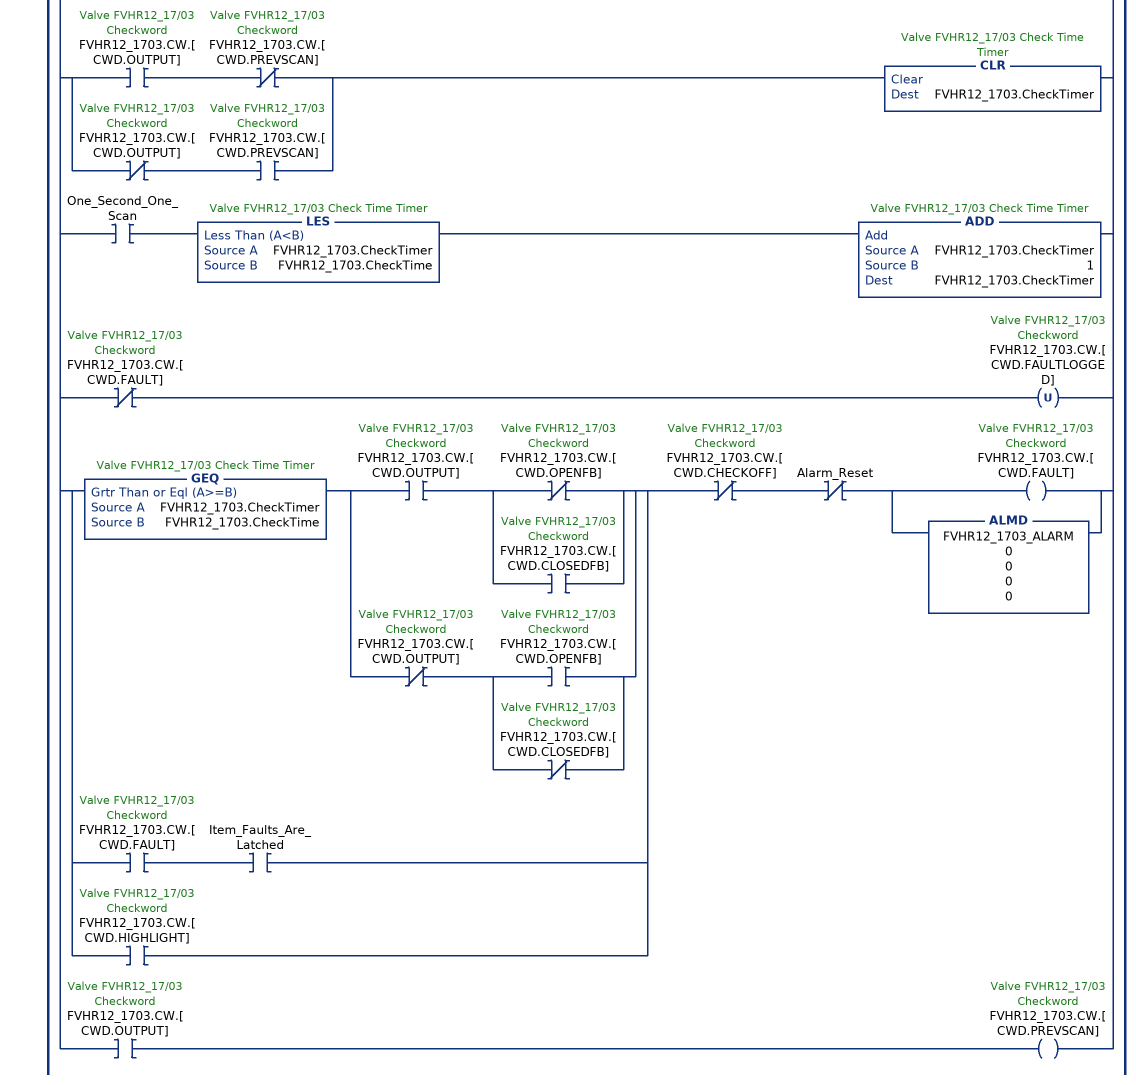
   71: [NEQ(FVHR12_1703.DriveBits,0) OTE(FVHR12_1703.CW.[CWD.AUTODRV]) ,[XIC(FVHR12_1703.CW.[CWD.AUTODRV]) XIO(FVHR12_1703.CW.[CWD.MANUAL]) ,XIC(FVHR12_1703.CW.[CWD.MANDRV]) XIC(FVHR12_1703.CW.[CWD.MANUAL]) ] OTE(FVHR12_1703.CW.[CWD.OUTPUT]) ,XIC(FVHR12_1703.CW.[CWD.OUTPUT]) OTE(FVHR12_1703_DR) ,XIC(S:FS) [OTU(FVHR12_1703.CW.[CWD.MANUAL]) ,LEQ(FVHR12_1703.CheckTime,0) MOV(Default_Check_Time,FVHR12_1703.CheckTime) ] ,[[XIC(FVHR12_1703_OP) XIO(Item_Simulation_Flag) ,XIC(Item_Simulation_Flag) XIC(FVHR12_1703.CW.[CWD.OUTPUT]) XIO(FVHR12_1703.CW.[CWD.SIMFAIL]) ] OTE(FVHR12_1703.CW.[CWD.OPENFB]) ,[XIC(FVHR12_1703_CL) XIO(Item_Simulation_Flag) ,XIC(Item_Simulation_Flag) XIO(FVHR12_1703.CW.[CWD.OUTPUT]) XIO(FVHR12_1703.CW.[CWD.SIMFAIL]) ] OTE(FVHR12_1703.CW.[CWD.CLOSEDFB]) ] ,[XIC(FVHR12_1703.CW.[CWD.OUTPUT]) XIO(FVHR12_1703.CW.[CWD.PREVSCAN]) ,XIO(FVHR12_1703.CW.[CWD.OUTPUT]) XIC(FVHR12_1703.CW.[CWD.PREVSCAN]) ] CLR(FVHR12_1703.CheckTimer) ,XIC(One_Second_One_Scan) LES(FVHR12_1703.CheckTimer,FVHR12_1703.CheckTime) ADD(FVHR12_1703.CheckTimer,1,FVHR12_1703.CheckTimer) ,XIO(FVHR12_1703.CW.[CWD.FAULT]) OTU(FVHR12_1703.CW.[CWD.FAULTLOGGED]) ,[GEQ(FVHR12_1703.CheckTimer,FVHR12_1703.CheckTime) [XIC(FVHR12_1703.CW.[CWD.OUTPUT]) [XIO(FVHR12_1703.CW.[CWD.OPENFB]) ,XIC(FVHR12_1703.CW.[CWD.CLOSEDFB]) ] ,XIO(FVHR12_1703.CW.[CWD.OUTPUT]) [XIC(FVHR12_1703.CW.[CWD.OPENFB]) ,XIO(FVHR12_1703.CW.[CWD.CLOSEDFB]) ] ] ,XIC(FVHR12_1703.CW.[CWD.FAULT]) XIC(Item_Faults_Are_Latched) ,XIC(FVHR12_1703.CW.[CWD.HIGHLIGHT]) ] XIO(FVHR12_1703.CW.[CWD.CHECKOFF]) XIO(Alarm_Reset) [OTE(FVHR12_1703.CW.[CWD.FAULT]) ,ALMD(FVHR12_1703_ALARM,0,0,0,0) ] ,XIC(FVHR12_1703.CW.[CWD.OUTPUT]) OTE(FVHR12_1703.CW.[CWD.PREVSCAN]) ];
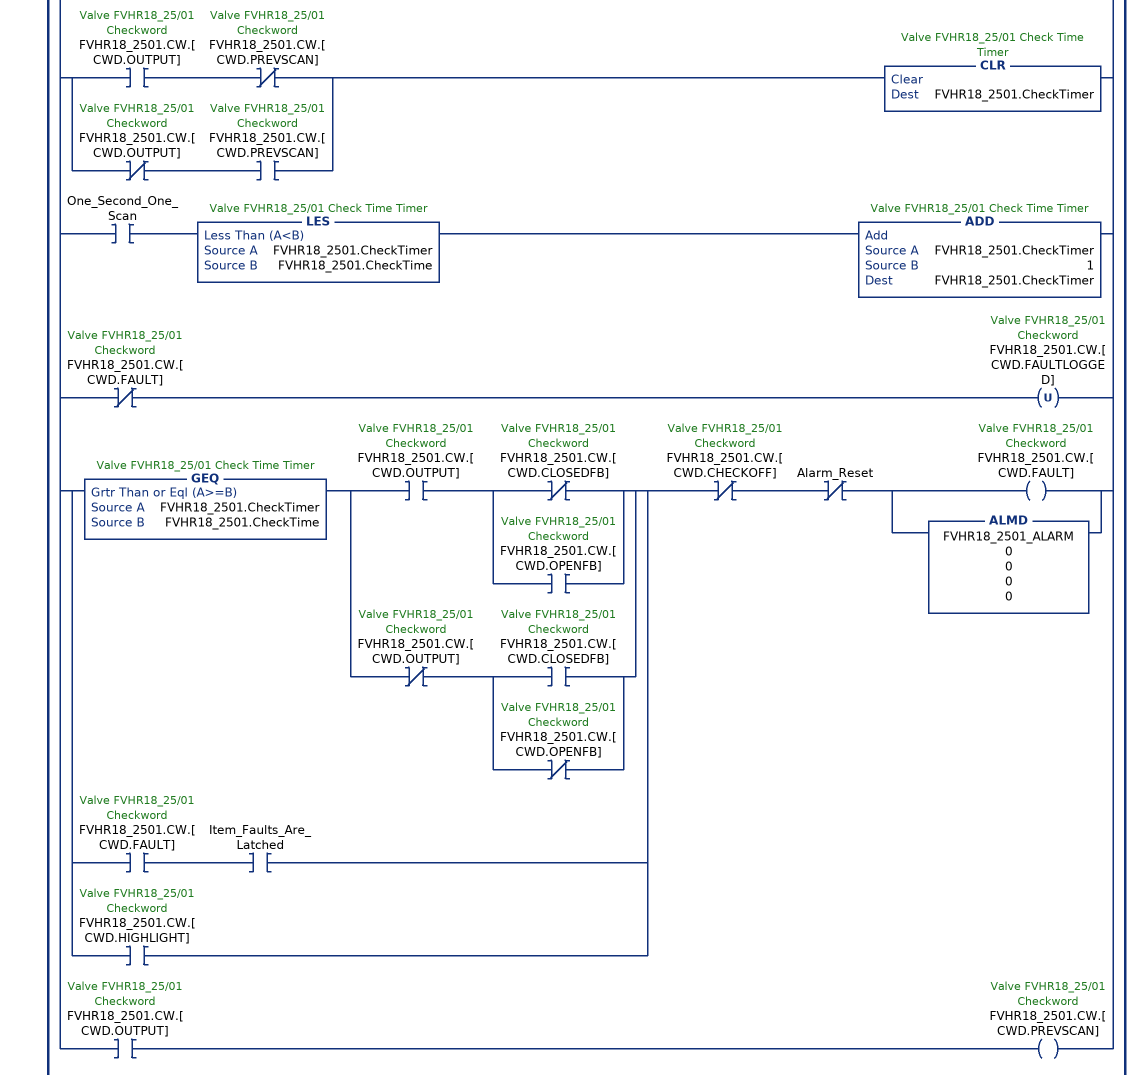
   72: [NEQ(FVHR18_2501.DriveBits,0) OTE(FVHR18_2501.CW.[CWD.AUTODRV]) ,[XIC(FVHR18_2501.CW.[CWD.AUTODRV]) XIO(FVHR18_2501.CW.[CWD.MANUAL]) ,XIC(FVHR18_2501.CW.[CWD.MANDRV]) XIC(FVHR18_2501.CW.[CWD.MANUAL]) ] OTE(FVHR18_2501.CW.[CWD.OUTPUT]) ,XIC(FVHR18_2501.CW.[CWD.OUTPUT]) OTE(FVHR18_2501_DR) ,XIC(S:FS) [OTU(FVHR18_2501.CW.[CWD.MANUAL]) ,LEQ(FVHR18_2501.CheckTime,0) MOV(Default_Check_Time,FVHR18_2501.CheckTime) ] ,[[XIC(FVHR18_2501_OP) XIO(Item_Simulation_Flag) ,XIC(Item_Simulation_Flag) XIC(FVHR18_2501.CW.[CWD.OUTPUT]) XIO(FVHR18_2501.CW.[CWD.SIMFAIL]) ] OTE(FVHR18_2501.CW.[CWD.OPENFB]) ,[XIC(FVHR18_2501_CL) XIO(Item_Simulation_Flag) ,XIC(Item_Simulation_Flag) XIO(FVHR18_2501.CW.[CWD.OUTPUT]) XIO(FVHR18_2501.CW.[CWD.SIMFAIL]) ] OTE(FVHR18_2501.CW.[CWD.CLOSEDFB]) ] ,[XIC(FVHR18_2501.CW.[CWD.OUTPUT]) XIO(FVHR18_2501.CW.[CWD.PREVSCAN]) ,XIO(FVHR18_2501.CW.[CWD.OUTPUT]) XIC(FVHR18_2501.CW.[CWD.PREVSCAN]) ] CLR(FVHR18_2501.CheckTimer) ,XIC(One_Second_One_Scan) LES(FVHR18_2501.CheckTimer,FVHR18_2501.CheckTime) ADD(FVHR18_2501.CheckTimer,1,FVHR18_2501.CheckTimer) ,XIO(FVHR18_2501.CW.[CWD.FAULT]) OTU(FVHR18_2501.CW.[CWD.FAULTLOGGED]) ,[GEQ(FVHR18_2501.CheckTimer,FVHR18_2501.CheckTime) [XIC(FVHR18_2501.CW.[CWD.OUTPUT]) [XIO(FVHR18_2501.CW.[CWD.CLOSEDFB]) ,XIC(FVHR18_2501.CW.[CWD.OPENFB]) ] ,XIO(FVHR18_2501.CW.[CWD.OUTPUT]) [XIC(FVHR18_2501.CW.[CWD.CLOSEDFB]) ,XIO(FVHR18_2501.CW.[CWD.OPENFB]) ] ] ,XIC(FVHR18_2501.CW.[CWD.FAULT]) XIC(Item_Faults_Are_Latched) ,XIC(FVHR18_2501.CW.[CWD.HIGHLIGHT]) ] XIO(FVHR18_2501.CW.[CWD.CHECKOFF]) XIO(Alarm_Reset) [OTE(FVHR18_2501.CW.[CWD.FAULT]) ,ALMD(FVHR18_2501_ALARM,0,0,0,0) ] ,XIC(FVHR18_2501.CW.[CWD.OUTPUT]) OTE(FVHR18_2501.CW.[CWD.PREVSCAN]) ];
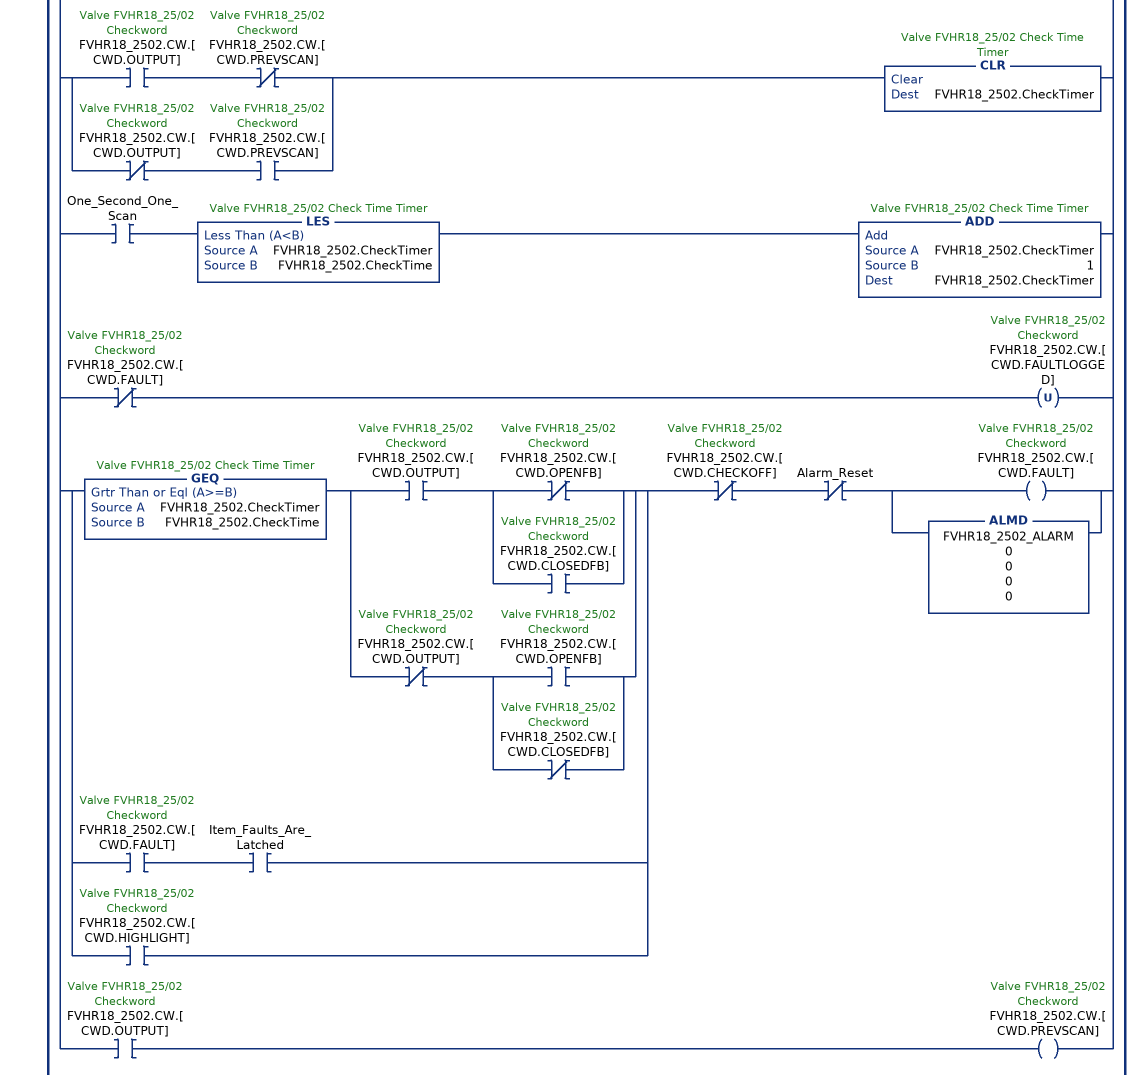
   73: [NEQ(FVHR18_2502.DriveBits,0) OTE(FVHR18_2502.CW.[CWD.AUTODRV]) ,[XIC(FVHR18_2502.CW.[CWD.AUTODRV]) XIO(FVHR18_2502.CW.[CWD.MANUAL]) ,XIC(FVHR18_2502.CW.[CWD.MANDRV]) XIC(FVHR18_2502.CW.[CWD.MANUAL]) ] OTE(FVHR18_2502.CW.[CWD.OUTPUT]) ,XIC(FVHR18_2502.CW.[CWD.OUTPUT]) OTE(FVHR18_2502_DR) ,XIC(S:FS) [OTU(FVHR18_2502.CW.[CWD.MANUAL]) ,LEQ(FVHR18_2502.CheckTime,0) MOV(Default_Check_Time,FVHR18_2502.CheckTime) ] ,[[XIC(FVHR18_2502_OP) XIO(Item_Simulation_Flag) ,XIC(Item_Simulation_Flag) XIC(FVHR18_2502.CW.[CWD.OUTPUT]) XIO(FVHR18_2502.CW.[CWD.SIMFAIL]) ] OTE(FVHR18_2502.CW.[CWD.OPENFB]) ,[XIC(FVHR18_2502_CL) XIO(Item_Simulation_Flag) ,XIC(Item_Simulation_Flag) XIO(FVHR18_2502.CW.[CWD.OUTPUT]) XIO(FVHR18_2502.CW.[CWD.SIMFAIL]) ] OTE(FVHR18_2502.CW.[CWD.CLOSEDFB]) ] ,[XIC(FVHR18_2502.CW.[CWD.OUTPUT]) XIO(FVHR18_2502.CW.[CWD.PREVSCAN]) ,XIO(FVHR18_2502.CW.[CWD.OUTPUT]) XIC(FVHR18_2502.CW.[CWD.PREVSCAN]) ] CLR(FVHR18_2502.CheckTimer) ,XIC(One_Second_One_Scan) LES(FVHR18_2502.CheckTimer,FVHR18_2502.CheckTime) ADD(FVHR18_2502.CheckTimer,1,FVHR18_2502.CheckTimer) ,XIO(FVHR18_2502.CW.[CWD.FAULT]) OTU(FVHR18_2502.CW.[CWD.FAULTLOGGED]) ,[GEQ(FVHR18_2502.CheckTimer,FVHR18_2502.CheckTime) [XIC(FVHR18_2502.CW.[CWD.OUTPUT]) [XIO(FVHR18_2502.CW.[CWD.OPENFB]) ,XIC(FVHR18_2502.CW.[CWD.CLOSEDFB]) ] ,XIO(FVHR18_2502.CW.[CWD.OUTPUT]) [XIC(FVHR18_2502.CW.[CWD.OPENFB]) ,XIO(FVHR18_2502.CW.[CWD.CLOSEDFB]) ] ] ,XIC(FVHR18_2502.CW.[CWD.FAULT]) XIC(Item_Faults_Are_Latched) ,XIC(FVHR18_2502.CW.[CWD.HIGHLIGHT]) ] XIO(FVHR18_2502.CW.[CWD.CHECKOFF]) XIO(Alarm_Reset) [OTE(FVHR18_2502.CW.[CWD.FAULT]) ,ALMD(FVHR18_2502_ALARM,0,0,0,0) ] ,XIC(FVHR18_2502.CW.[CWD.OUTPUT]) OTE(FVHR18_2502.CW.[CWD.PREVSCAN]) ];
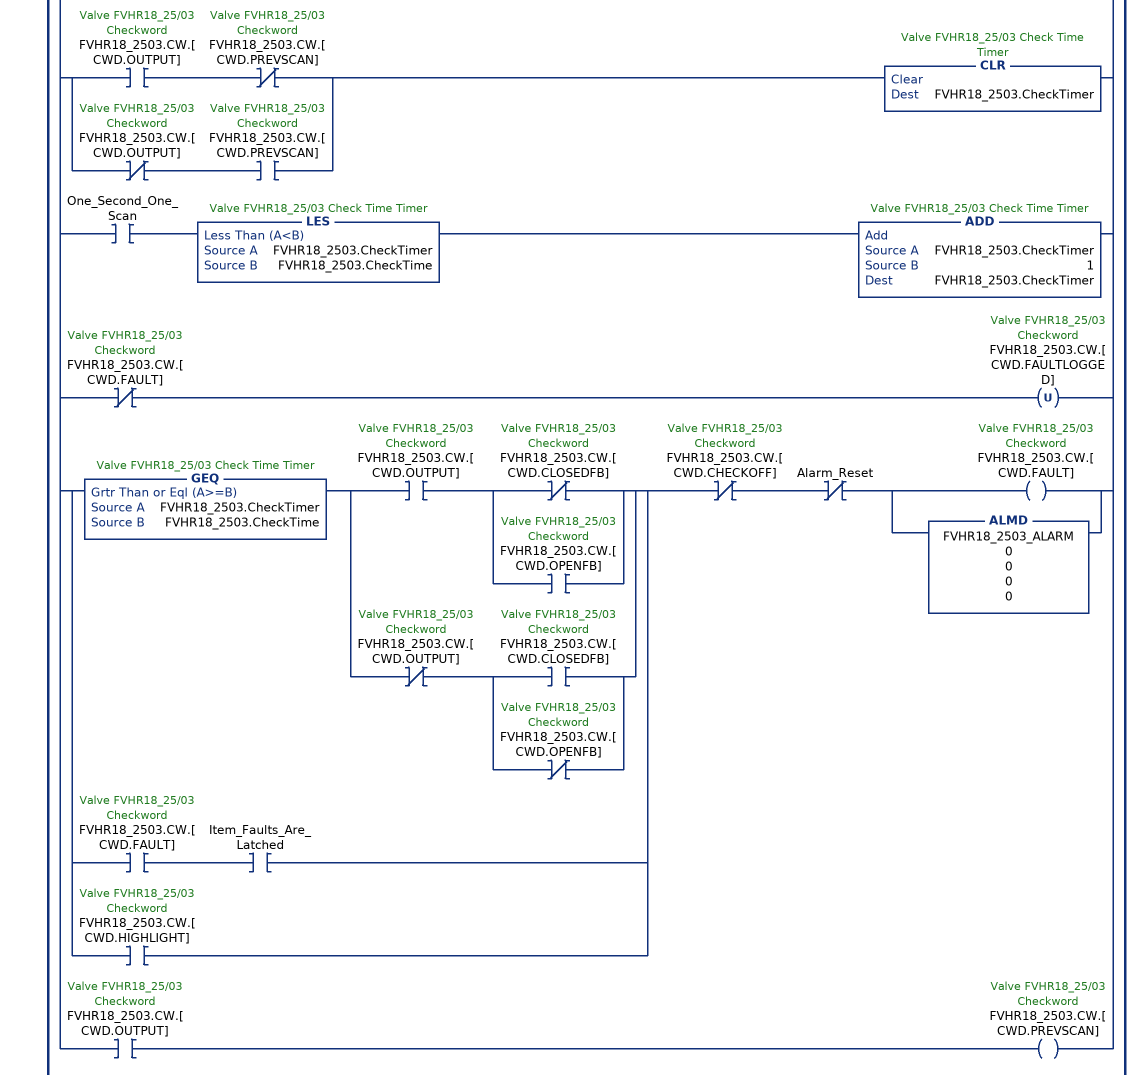
   74: [NEQ(FVHR18_2503.DriveBits,0) OTE(FVHR18_2503.CW.[CWD.AUTODRV]) ,[XIC(FVHR18_2503.CW.[CWD.AUTODRV]) XIO(FVHR18_2503.CW.[CWD.MANUAL]) ,XIC(FVHR18_2503.CW.[CWD.MANDRV]) XIC(FVHR18_2503.CW.[CWD.MANUAL]) ] OTE(FVHR18_2503.CW.[CWD.OUTPUT]) ,XIC(FVHR18_2503.CW.[CWD.OUTPUT]) OTE(FVHR18_2503_DR) ,XIC(S:FS) [OTU(FVHR18_2503.CW.[CWD.MANUAL]) ,LEQ(FVHR18_2503.CheckTime,0) MOV(Default_Check_Time,FVHR18_2503.CheckTime) ] ,[[XIC(FVHR18_2503_OP) XIO(Item_Simulation_Flag) ,XIC(Item_Simulation_Flag) XIC(FVHR18_2503.CW.[CWD.OUTPUT]) XIO(FVHR18_2503.CW.[CWD.SIMFAIL]) ] OTE(FVHR18_2503.CW.[CWD.OPENFB]) ,[XIC(FVHR18_2503_CL) XIO(Item_Simulation_Flag) ,XIC(Item_Simulation_Flag) XIO(FVHR18_2503.CW.[CWD.OUTPUT]) XIO(FVHR18_2503.CW.[CWD.SIMFAIL]) ] OTE(FVHR18_2503.CW.[CWD.CLOSEDFB]) ] ,[XIC(FVHR18_2503.CW.[CWD.OUTPUT]) XIO(FVHR18_2503.CW.[CWD.PREVSCAN]) ,XIO(FVHR18_2503.CW.[CWD.OUTPUT]) XIC(FVHR18_2503.CW.[CWD.PREVSCAN]) ] CLR(FVHR18_2503.CheckTimer) ,XIC(One_Second_One_Scan) LES(FVHR18_2503.CheckTimer,FVHR18_2503.CheckTime) ADD(FVHR18_2503.CheckTimer,1,FVHR18_2503.CheckTimer) ,XIO(FVHR18_2503.CW.[CWD.FAULT]) OTU(FVHR18_2503.CW.[CWD.FAULTLOGGED]) ,[GEQ(FVHR18_2503.CheckTimer,FVHR18_2503.CheckTime) [XIC(FVHR18_2503.CW.[CWD.OUTPUT]) [XIO(FVHR18_2503.CW.[CWD.CLOSEDFB]) ,XIC(FVHR18_2503.CW.[CWD.OPENFB]) ] ,XIO(FVHR18_2503.CW.[CWD.OUTPUT]) [XIC(FVHR18_2503.CW.[CWD.CLOSEDFB]) ,XIO(FVHR18_2503.CW.[CWD.OPENFB]) ] ] ,XIC(FVHR18_2503.CW.[CWD.FAULT]) XIC(Item_Faults_Are_Latched) ,XIC(FVHR18_2503.CW.[CWD.HIGHLIGHT]) ] XIO(FVHR18_2503.CW.[CWD.CHECKOFF]) XIO(Alarm_Reset) [OTE(FVHR18_2503.CW.[CWD.FAULT]) ,ALMD(FVHR18_2503_ALARM,0,0,0,0) ] ,XIC(FVHR18_2503.CW.[CWD.OUTPUT]) OTE(FVHR18_2503.CW.[CWD.PREVSCAN]) ];
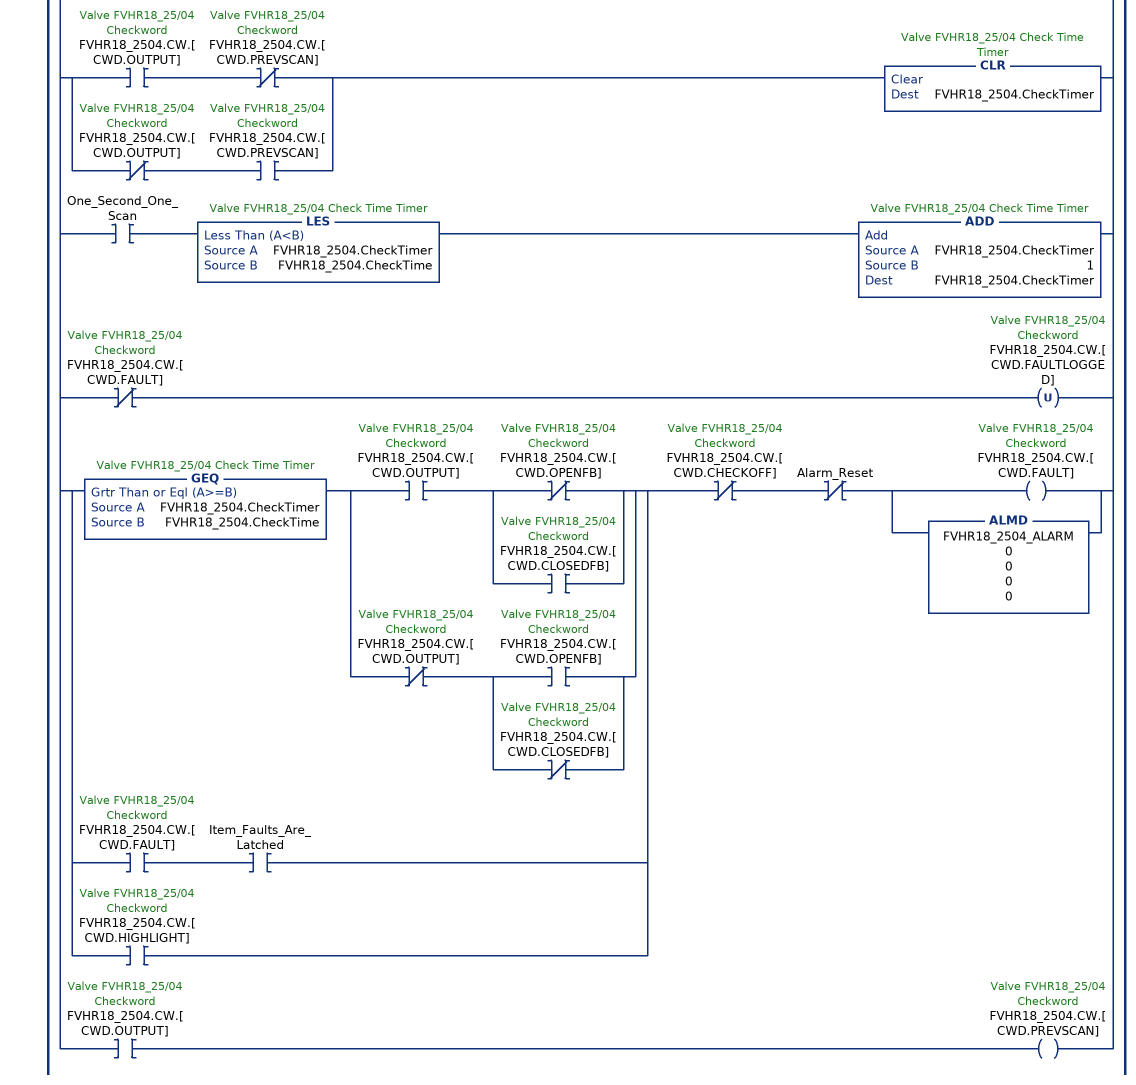
   75: [NEQ(FVHR18_2504.DriveBits,0) OTE(FVHR18_2504.CW.[CWD.AUTODRV]) ,[XIC(FVHR18_2504.CW.[CWD.AUTODRV]) XIO(FVHR18_2504.CW.[CWD.MANUAL]) ,XIC(FVHR18_2504.CW.[CWD.MANDRV]) XIC(FVHR18_2504.CW.[CWD.MANUAL]) ] OTE(FVHR18_2504.CW.[CWD.OUTPUT]) ,XIC(FVHR18_2504.CW.[CWD.OUTPUT]) OTE(FVHR18_2504_DR) ,XIC(S:FS) [OTU(FVHR18_2504.CW.[CWD.MANUAL]) ,LEQ(FVHR18_2504.CheckTime,0) MOV(Default_Check_Time,FVHR18_2504.CheckTime) ] ,[[XIC(FVHR18_2504_OP) XIO(Item_Simulation_Flag) ,XIC(Item_Simulation_Flag) XIC(FVHR18_2504.CW.[CWD.OUTPUT]) XIO(FVHR18_2504.CW.[CWD.SIMFAIL]) ] OTE(FVHR18_2504.CW.[CWD.OPENFB]) ,[XIC(FVHR18_2504_CL) XIO(Item_Simulation_Flag) ,XIC(Item_Simulation_Flag) XIO(FVHR18_2504.CW.[CWD.OUTPUT]) XIO(FVHR18_2504.CW.[CWD.SIMFAIL]) ] OTE(FVHR18_2504.CW.[CWD.CLOSEDFB]) ] ,[XIC(FVHR18_2504.CW.[CWD.OUTPUT]) XIO(FVHR18_2504.CW.[CWD.PREVSCAN]) ,XIO(FVHR18_2504.CW.[CWD.OUTPUT]) XIC(FVHR18_2504.CW.[CWD.PREVSCAN]) ] CLR(FVHR18_2504.CheckTimer) ,XIC(One_Second_One_Scan) LES(FVHR18_2504.CheckTimer,FVHR18_2504.CheckTime) ADD(FVHR18_2504.CheckTimer,1,FVHR18_2504.CheckTimer) ,XIO(FVHR18_2504.CW.[CWD.FAULT]) OTU(FVHR18_2504.CW.[CWD.FAULTLOGGED]) ,[GEQ(FVHR18_2504.CheckTimer,FVHR18_2504.CheckTime) [XIC(FVHR18_2504.CW.[CWD.OUTPUT]) [XIO(FVHR18_2504.CW.[CWD.OPENFB]) ,XIC(FVHR18_2504.CW.[CWD.CLOSEDFB]) ] ,XIO(FVHR18_2504.CW.[CWD.OUTPUT]) [XIC(FVHR18_2504.CW.[CWD.OPENFB]) ,XIO(FVHR18_2504.CW.[CWD.CLOSEDFB]) ] ] ,XIC(FVHR18_2504.CW.[CWD.FAULT]) XIC(Item_Faults_Are_Latched) ,XIC(FVHR18_2504.CW.[CWD.HIGHLIGHT]) ] XIO(FVHR18_2504.CW.[CWD.CHECKOFF]) XIO(Alarm_Reset) [OTE(FVHR18_2504.CW.[CWD.FAULT]) ,ALMD(FVHR18_2504_ALARM,0,0,0,0) ] ,XIC(FVHR18_2504.CW.[CWD.OUTPUT]) OTE(FVHR18_2504.CW.[CWD.PREVSCAN]) ];
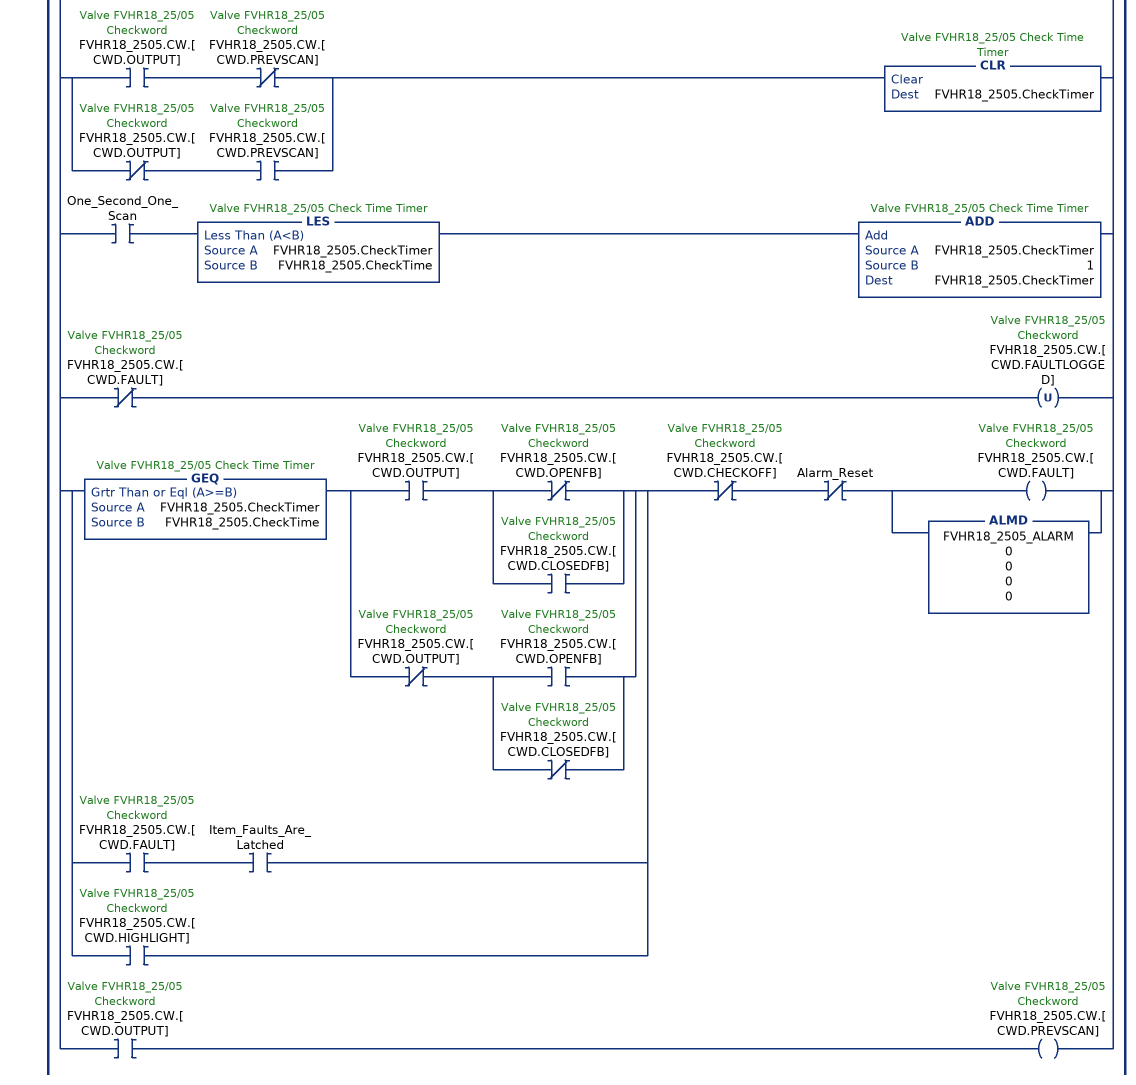
   76: [NEQ(FVHR18_2505.DriveBits,0) OTE(FVHR18_2505.CW.[CWD.AUTODRV]) ,[XIC(FVHR18_2505.CW.[CWD.AUTODRV]) XIO(FVHR18_2505.CW.[CWD.MANUAL]) ,XIC(FVHR18_2505.CW.[CWD.MANDRV]) XIC(FVHR18_2505.CW.[CWD.MANUAL]) ] OTE(FVHR18_2505.CW.[CWD.OUTPUT]) ,XIC(FVHR18_2505.CW.[CWD.OUTPUT]) OTE(FVHR18_2505_DR) ,XIC(S:FS) [OTU(FVHR18_2505.CW.[CWD.MANUAL]) ,LEQ(FVHR18_2505.CheckTime,0) MOV(Default_Check_Time,FVHR18_2505.CheckTime) ] ,[[XIC(FVHR18_2505_OP) XIO(Item_Simulation_Flag) ,XIC(Item_Simulation_Flag) XIC(FVHR18_2505.CW.[CWD.OUTPUT]) XIO(FVHR18_2505.CW.[CWD.SIMFAIL]) ] OTE(FVHR18_2505.CW.[CWD.OPENFB]) ,[XIC(FVHR18_2505_CL) XIO(Item_Simulation_Flag) ,XIC(Item_Simulation_Flag) XIO(FVHR18_2505.CW.[CWD.OUTPUT]) XIO(FVHR18_2505.CW.[CWD.SIMFAIL]) ] OTE(FVHR18_2505.CW.[CWD.CLOSEDFB]) ] ,[XIC(FVHR18_2505.CW.[CWD.OUTPUT]) XIO(FVHR18_2505.CW.[CWD.PREVSCAN]) ,XIO(FVHR18_2505.CW.[CWD.OUTPUT]) XIC(FVHR18_2505.CW.[CWD.PREVSCAN]) ] CLR(FVHR18_2505.CheckTimer) ,XIC(One_Second_One_Scan) LES(FVHR18_2505.CheckTimer,FVHR18_2505.CheckTime) ADD(FVHR18_2505.CheckTimer,1,FVHR18_2505.CheckTimer) ,XIO(FVHR18_2505.CW.[CWD.FAULT]) OTU(FVHR18_2505.CW.[CWD.FAULTLOGGED]) ,[GEQ(FVHR18_2505.CheckTimer,FVHR18_2505.CheckTime) [XIC(FVHR18_2505.CW.[CWD.OUTPUT]) [XIO(FVHR18_2505.CW.[CWD.OPENFB]) ,XIC(FVHR18_2505.CW.[CWD.CLOSEDFB]) ] ,XIO(FVHR18_2505.CW.[CWD.OUTPUT]) [XIC(FVHR18_2505.CW.[CWD.OPENFB]) ,XIO(FVHR18_2505.CW.[CWD.CLOSEDFB]) ] ] ,XIC(FVHR18_2505.CW.[CWD.FAULT]) XIC(Item_Faults_Are_Latched) ,XIC(FVHR18_2505.CW.[CWD.HIGHLIGHT]) ] XIO(FVHR18_2505.CW.[CWD.CHECKOFF]) XIO(Alarm_Reset) [OTE(FVHR18_2505.CW.[CWD.FAULT]) ,ALMD(FVHR18_2505_ALARM,0,0,0,0) ] ,XIC(FVHR18_2505.CW.[CWD.OUTPUT]) OTE(FVHR18_2505.CW.[CWD.PREVSCAN]) ];
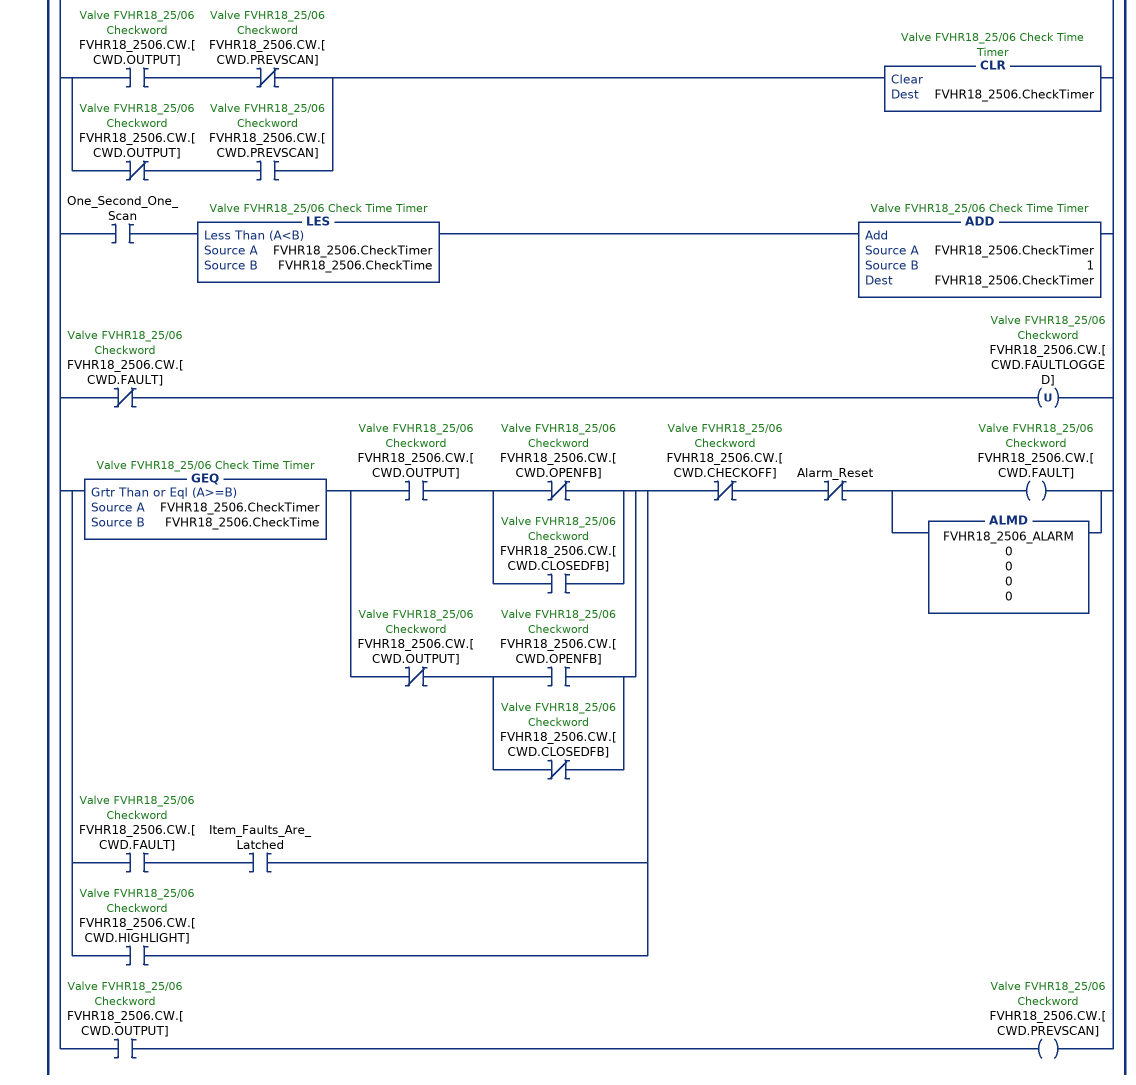
   77: [NEQ(FVHR18_2506.DriveBits,0) OTE(FVHR18_2506.CW.[CWD.AUTODRV]) ,[XIC(FVHR18_2506.CW.[CWD.AUTODRV]) XIO(FVHR18_2506.CW.[CWD.MANUAL]) ,XIC(FVHR18_2506.CW.[CWD.MANDRV]) XIC(FVHR18_2506.CW.[CWD.MANUAL]) ] OTE(FVHR18_2506.CW.[CWD.OUTPUT]) ,XIC(FVHR18_2506.CW.[CWD.OUTPUT]) OTE(FVHR18_2506_DR) ,XIC(S:FS) [OTU(FVHR18_2506.CW.[CWD.MANUAL]) ,LEQ(FVHR18_2506.CheckTime,0) MOV(Default_Check_Time,FVHR18_2506.CheckTime) ] ,[[XIC(FVHR18_2506_OP) XIO(Item_Simulation_Flag) ,XIC(Item_Simulation_Flag) XIC(FVHR18_2506.CW.[CWD.OUTPUT]) XIO(FVHR18_2506.CW.[CWD.SIMFAIL]) ] OTE(FVHR18_2506.CW.[CWD.OPENFB]) ,[XIC(FVHR18_2506_CL) XIO(Item_Simulation_Flag) ,XIC(Item_Simulation_Flag) XIO(FVHR18_2506.CW.[CWD.OUTPUT]) XIO(FVHR18_2506.CW.[CWD.SIMFAIL]) ] OTE(FVHR18_2506.CW.[CWD.CLOSEDFB]) ] ,[XIC(FVHR18_2506.CW.[CWD.OUTPUT]) XIO(FVHR18_2506.CW.[CWD.PREVSCAN]) ,XIO(FVHR18_2506.CW.[CWD.OUTPUT]) XIC(FVHR18_2506.CW.[CWD.PREVSCAN]) ] CLR(FVHR18_2506.CheckTimer) ,XIC(One_Second_One_Scan) LES(FVHR18_2506.CheckTimer,FVHR18_2506.CheckTime) ADD(FVHR18_2506.CheckTimer,1,FVHR18_2506.CheckTimer) ,XIO(FVHR18_2506.CW.[CWD.FAULT]) OTU(FVHR18_2506.CW.[CWD.FAULTLOGGED]) ,[GEQ(FVHR18_2506.CheckTimer,FVHR18_2506.CheckTime) [XIC(FVHR18_2506.CW.[CWD.OUTPUT]) [XIO(FVHR18_2506.CW.[CWD.OPENFB]) ,XIC(FVHR18_2506.CW.[CWD.CLOSEDFB]) ] ,XIO(FVHR18_2506.CW.[CWD.OUTPUT]) [XIC(FVHR18_2506.CW.[CWD.OPENFB]) ,XIO(FVHR18_2506.CW.[CWD.CLOSEDFB]) ] ] ,XIC(FVHR18_2506.CW.[CWD.FAULT]) XIC(Item_Faults_Are_Latched) ,XIC(FVHR18_2506.CW.[CWD.HIGHLIGHT]) ] XIO(FVHR18_2506.CW.[CWD.CHECKOFF]) XIO(Alarm_Reset) [OTE(FVHR18_2506.CW.[CWD.FAULT]) ,ALMD(FVHR18_2506_ALARM,0,0,0,0) ] ,XIC(FVHR18_2506.CW.[CWD.OUTPUT]) OTE(FVHR18_2506.CW.[CWD.PREVSCAN]) ];
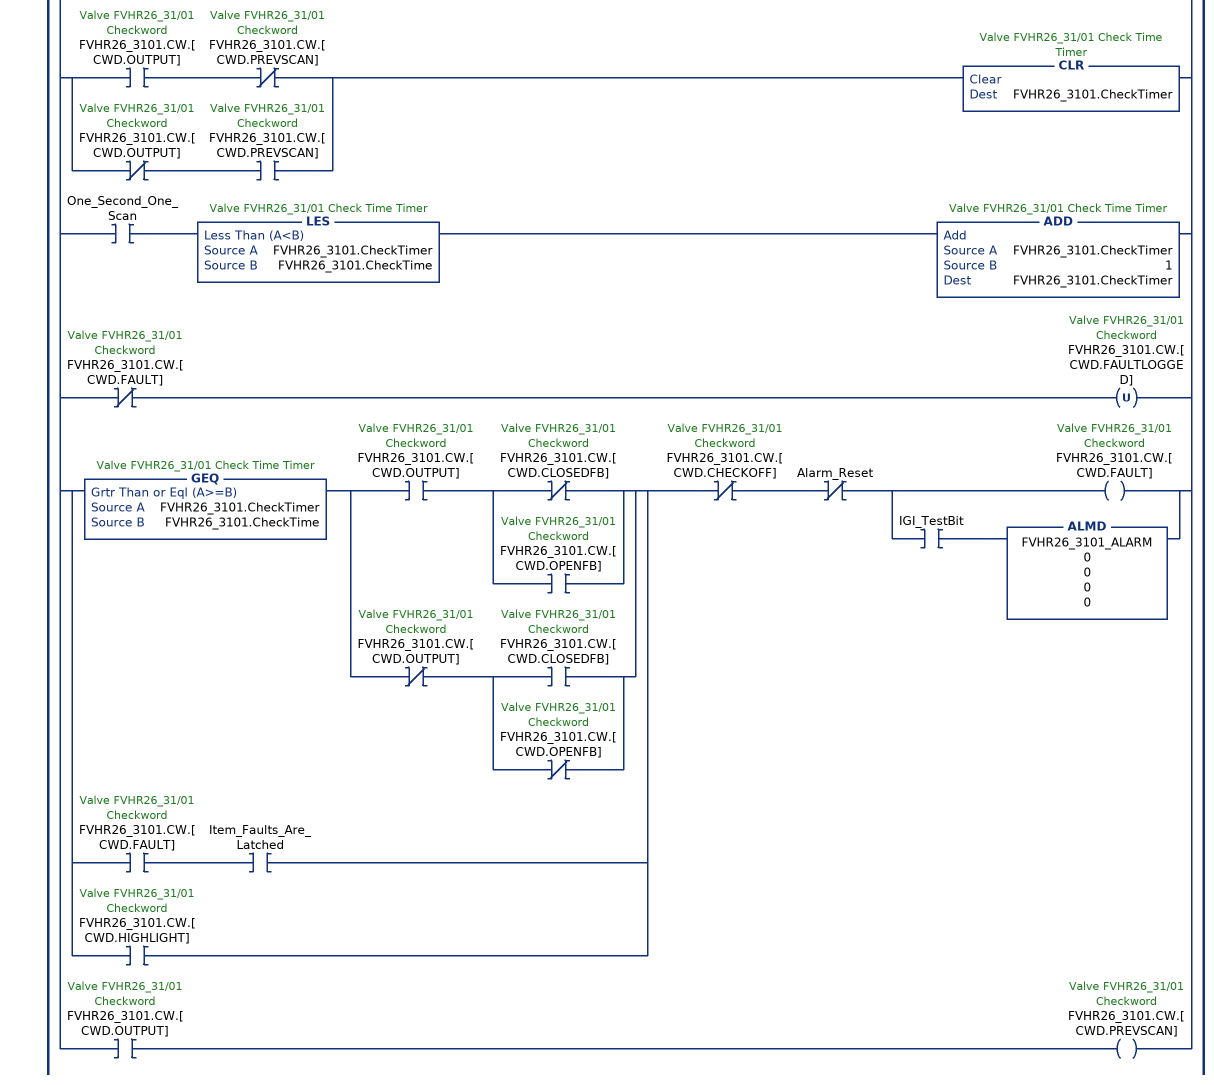
   78: [NEQ(FVHR26_3101.DriveBits,0) OTE(FVHR26_3101.CW.[CWD.AUTODRV]) ,[XIC(FVHR26_3101.CW.[CWD.AUTODRV]) XIO(FVHR26_3101.CW.[CWD.MANUAL]) ,XIC(FVHR26_3101.CW.[CWD.MANDRV]) XIC(FVHR26_3101.CW.[CWD.MANUAL]) ] OTE(FVHR26_3101.CW.[CWD.OUTPUT]) ,XIC(FVHR26_3101.CW.[CWD.OUTPUT]) OTE(FVHR26_3101_DR) ,XIC(S:FS) [OTU(FVHR26_3101.CW.[CWD.MANUAL]) ,LEQ(FVHR26_3101.CheckTime,0) MOV(Default_Check_Time,FVHR26_3101.CheckTime) ] ,[[XIC(FVHR26_3101_OP) XIO(Item_Simulation_Flag) ,XIC(Item_Simulation_Flag) XIC(FVHR26_3101.CW.[CWD.OUTPUT]) XIO(FVHR26_3101.CW.[CWD.SIMFAIL]) ] OTE(FVHR26_3101.CW.[CWD.OPENFB]) ,[XIC(FVHR26_3101_CL) XIO(Item_Simulation_Flag) ,XIC(Item_Simulation_Flag) XIO(FVHR26_3101.CW.[CWD.OUTPUT]) XIO(FVHR26_3101.CW.[CWD.SIMFAIL]) ] OTE(FVHR26_3101.CW.[CWD.CLOSEDFB]) ] ,[XIC(FVHR26_3101.CW.[CWD.OUTPUT]) XIO(FVHR26_3101.CW.[CWD.PREVSCAN]) ,XIO(FVHR26_3101.CW.[CWD.OUTPUT]) XIC(FVHR26_3101.CW.[CWD.PREVSCAN]) ] CLR(FVHR26_3101.CheckTimer) ,XIC(One_Second_One_Scan) LES(FVHR26_3101.CheckTimer,FVHR26_3101.CheckTime) ADD(FVHR26_3101.CheckTimer,1,FVHR26_3101.CheckTimer) ,XIO(FVHR26_3101.CW.[CWD.FAULT]) OTU(FVHR26_3101.CW.[CWD.FAULTLOGGED]) ,[GEQ(FVHR26_3101.CheckTimer,FVHR26_3101.CheckTime) [XIC(FVHR26_3101.CW.[CWD.OUTPUT]) [XIO(FVHR26_3101.CW.[CWD.CLOSEDFB]) ,XIC(FVHR26_3101.CW.[CWD.OPENFB]) ] ,XIO(FVHR26_3101.CW.[CWD.OUTPUT]) [XIC(FVHR26_3101.CW.[CWD.CLOSEDFB]) ,XIO(FVHR26_3101.CW.[CWD.OPENFB]) ] ] ,XIC(FVHR26_3101.CW.[CWD.FAULT]) XIC(Item_Faults_Are_Latched) ,XIC(FVHR26_3101.CW.[CWD.HIGHLIGHT]) ] XIO(FVHR26_3101.CW.[CWD.CHECKOFF]) XIO(Alarm_Reset) [OTE(FVHR26_3101.CW.[CWD.FAULT]) ,XIC(IGI_TestBit) ALMD(FVHR26_3101_ALARM,0,0,0,0) ] ,XIC(FVHR26_3101.CW.[CWD.OUTPUT]) OTE(FVHR26_3101.CW.[CWD.PREVSCAN]) ];
